VERSION : 0.1
   VAR
      _1s1 : Bool;
      _1s2 : Bool;
      _1s3 : Bool;
      _1s4 : Bool;
      _1s5 : Bool;
      _1s6 : Bool;
      _1s7 : Bool;
      _1s8 : Bool;
      _1s9 : Bool;
      _1s10 : Bool;
      _1sReserva2 : Bool;
      _1sReserva3 : Bool;
      _1sReserva4 : Bool;
      _1sReserva5 : Bool;
      _1sReserva6 : Bool;
      _1sReserva7 : Bool;
      _2s1 : Bool;
      _2s2 : Bool;
      _2s3 : Bool;
      _2s4 : Bool;
      _2s5 : Bool;
      _2s6 : Bool;
      _2s7 : Bool;
      _2s8 : Bool;
      _2s9 : Bool;
      _2s10 : Bool;
      _2sReserva2 : Bool;
      _2sReserva3 : Bool;
      _2sReserva4 : Bool;
      _2sReserva5 : Bool;
      _2sReserva6 : Bool;
      _2sReserva7 : Bool;
      _3s1 : Bool;
      _3s2 : Bool;
      _3s3 : Bool;
      _3s4 : Bool;
      _3s5 : Bool;
      _3s6 : Bool;
      _3s7 : Bool;
      _3s8 : Bool;
      _3s9 : Bool;
      _3s10 : Bool;
      _3Reserva2 : Bool;
      _3Reserva3 : Bool;
      _3Reserva4 : Bool;
      _3Reserva5 : Bool;
      _3Reserva6 : Bool;
      _3Reserva7 : Bool;
      _4s1 : Bool;
      _4s2 : Bool;
      _4s3 : Bool;
      _4s4 : Bool;
      _4s5 : Bool;
      _4s6 : Bool;
      _4s7 : Bool;
      _4s8 : Bool;
      _4s9 : Bool;
      _4s10 : Bool;
      _4sReserva2 : Bool;
      _4sReserva3 : Bool;
      _4sReserva4 : Bool;
      _4sReserva5 : Bool;
      _4sReserva6 : Bool;
      _4sReserva7 : Bool;
      _5s1 : Bool;
      _5s2 : Bool;
      _5s3 : Bool;
      _5s4 : Bool;
      _5s5 : Bool;
      _5s6 : Bool;
      _5s7 : Bool;
      _5s8 : Bool;
      _5s9 : Bool;
      _5s10 : Bool;
      _5sReserva2 : Bool;
      _5sReserva3 : Bool;
      _5sReserva4 : Bool;
      _5sReserva5 : Bool;
      _5sReserva6 : Bool;
      _5sReserva7 : Bool;
      _6s1 : Bool;
      _6s2 : Bool;
      _6s3 : Bool;
      _6s4 : Bool;
      _6s5 : Bool;
      _6s6 : Bool;
      _6s7 : Bool;
      _6s8 : Bool;
      _6s9 : Bool;
      _6s10 : Bool;
      _6sReserva2 : Bool;
      _6sReserva3 : Bool;
      _6sReserva4 : Bool;
      _6sReserva5 : Bool;
      _6sReserva6 : Bool;
      _6sReserva7 : Bool;
      _0s1 : Bool;   // No requiere Compresores
      _0s2 : Bool;   // Requiere 1 Compresor
      _0s3 : Bool;   // Requiere 2 Compresores
      _0s4 : Bool;   // Requiere 3 Compresores
      _0s5 : Bool;   // Requiere 4 Compresores
      _0s6 : Bool;   // Requiere 5 Compresores
      _0s7 : Bool;
      _0s8 : Bool;
      _0s9 : Bool;
      _0s10 : Bool;
      _0sReserva2 : Bool;
      _0sReserva3 : Bool;
      _0sReserva4 : Bool;
      _0sReserva5 : Bool;
      _0sReserva6 : Bool;
      _0sReserva7 : Bool;
   END_VAR
BEGIN
END_DATA_BLOCK

DATA_BLOCK "Concatenadoras"   // DB127
{ S7_Optimized_Access := 'FALSE' }
VERSION : 0.1
   VAR
      _1c1 : Bool;
      _1c2 : Bool;
      _1c3 : Bool;
      _1c4 : Bool;
      _1c5 : Bool;
      _1c6 : Bool;
      _1c7 : Bool;
      _1c8 : Bool;
      _1c9 : Bool;
      _1c10 : Bool;
      _1cReserva2 : Bool;
      _1cReserva3 : Bool;
      _1cReserva4 : Bool;
      _1cReserva5 : Bool;
      _1cReserva6 : Bool;
      _1cReserva7 : Bool;
      _2c1 : Bool;
      _2c2 : Bool;
      _2c3 : Bool;
      _2c4 : Bool;
      _2c5 : Bool;
      _2c6 : Bool;
      _2c7 : Bool;
      _2c8 : Bool;
      _2c9 : Bool;
      _2c10 : Bool;
      _2cReserva2 : Bool;
      _2cReserva3 : Bool;
      _2cReserva4 : Bool;
      _2cReserva5 : Bool;
      _2cReserva6 : Bool;
      _2cReserva7 : Bool;
      _3c1 : Bool;
      _3c2 : Bool;
      _3c3 : Bool;
      _3c4 : Bool;
      _3c5 : Bool;
      _3c6 : Bool;
      _3c7 : Bool;
      _3c8 : Bool;
      _3c9 : Bool;
      _3c10 : Bool;
      _3cReserva2 : Bool;
      _3cReserva3 : Bool;
      _3cReserva4 : Bool;
      _3cReserva5 : Bool;
      _3cReserva6 : Bool;
      _3cReserva7 : Bool;
      _4c1 : Bool;
      _4c2 : Bool;
      _4c3 : Bool;
      _4c4 : Bool;
      _4c5 : Bool;
      _4c6 : Bool;
      _4c7 : Bool;
      _4c8 : Bool;
      _4c9 : Bool;
      _4c10 : Bool;
      _4cReserva2 : Bool;
      _4cReserva3 : Bool;
      _4cReserva4 : Bool;
      _4cReserva5 : Bool;
      _4cReserva6 : Bool;
      _4cReserva7 : Bool;
      _5c1 : Bool;
      _5c2 : Bool;
      _5c3 : Bool;
      _5c4 : Bool;
      _5c5 : Bool;
      _5c6 : Bool;
      _5c7 : Bool;
      _5c8 : Bool;
      _5c9 : Bool;
      _5c10 : Bool;
      _5cReserva2 : Bool;
      _5cReserva3 : Bool;
      _5cReserva4 : Bool;
      _5cReserva5 : Bool;
      _5cReserva6 : Bool;
      _5cReserva7 : Bool;
      _6c1 : Bool;
      _6c2 : Bool;
      _6c3 : Bool;
      _6c4 : Bool;
      _6c5 : Bool;
      _6c6 : Bool;
      _6c7 : Bool;
      _6c8 : Bool;
      _6c9 : Bool;
      _6c10 : Bool;
      _6cReserva2 : Bool;
      _6cReserva3 : Bool;
      _6cReserva4 : Bool;
      _6cReserva5 : Bool;
      _6cReserva6 : Bool;
      _6cReserva7 : Bool;
      _0c1 : Bool;   // No requiere Compresores
      _0c2 : Bool;   // Requiere 1 Compresor
      _0c3 : Bool;   // Requiere 2 Compresores
      _0c4 : Bool;   // Requiere 3 Compresores
      _0c5 : Bool;   // Requiere 4 Compresores
      _0c6 : Bool;   // Requiere 5 Compresores
      _0c7 : Bool;
      _0c8 : Bool;
      _0c9 : Bool;
      _0c10 : Bool;
      _0cReserva2 : Bool;
      _0cReserva3 : Bool;
      _0cReserva4 : Bool;
      _0cReserva5 : Bool;
      _0cReserva6 : Bool;
      _0cReserva7 : Bool;
   END_VAR
BEGIN
END_DATA_BLOCK

DATA_BLOCK "Prioritarias"   // DB128
{ S7_Optimized_Access := 'FALSE' }
VERSION : 0.1
   VAR
      _1p1 : Bool;
      _1p2 : Bool;
      _1p3 : Bool;
      _1p4 : Bool;
      _1p5 : Bool;
      _1p6 : Bool;
      _1p7 : Bool;
      _1p8 : Bool;
      _1p9 : Bool;
      _1p10 : Bool;
      _1pReserva2 : Bool;
      _1pReserva3 : Bool;
      _1pReserva4 : Bool;
      _1pReserva5 : Bool;
      _1pReserva6 : Bool;
      _1pReserva7 : Bool;
      _2p1 : Bool;
      _2p2 : Bool;
      _2p3 : Bool;
      _2p4 : Bool;
      _2p5 : Bool;
      _2p6 : Bool;
      _2p7 : Bool;
      _2p8 : Bool;
      _2p9 : Bool;
      _2p10 : Bool;
      _2pReserva2 : Bool;
      _2pReserva3 : Bool;
      _2pReserva4 : Bool;
      _2pReserva5 : Bool;
      _2pReserva6 : Bool;
      _2pReserva7 : Bool;
      _3p1 : Bool;
      _3p2 : Bool;
      _3p3 : Bool;
      _3p4 : Bool;
      _3p5 : Bool;
      _3p6 : Bool;
      _3p7 : Bool;
      _3p8 : Bool;
      _3p9 : Bool;
      _3p10 : Bool;
      _3pReserva2 : Bool;
      _3pReserva3 : Bool;
      _3pReserva4 : Bool;
      _3pReserva5 : Bool;
      _3pReserva6 : Bool;
      _3pReserva7 : Bool;
      _4p1 : Bool;
      _4p2 : Bool;
      _4p3 : Bool;
      _4p4 : Bool;
      _4p5 : Bool;
      _4p6 : Bool;
      _4p7 : Bool;
      _4p8 : Bool;
      _4p9 : Bool;
      _4p10 : Bool;
      _4pReserva2 : Bool;
      _4pReserva3 : Bool;
      _4pReserva4 : Bool;
      _4pReserva5 : Bool;
      _4pReserva6 : Bool;
      _4pReserva7 : Bool;
      _5p1 : Bool;
      _5p2 : Bool;
      _5p3 : Bool;
      _5p4 : Bool;
      _5p5 : Bool;
      _5p6 : Bool;
      _5p7 : Bool;
      _5p8 : Bool;
      _5p9 : Bool;
      _5p10 : Bool;
      _5pReserva2 : Bool;
      _5pReserva3 : Bool;
      _5pReserva4 : Bool;
      _5pReserva5 : Bool;
      _5pReserva6 : Bool;
      _5pReserva7 : Bool;
      _6p1 : Bool;
      _6p2 : Bool;
      _6p3 : Bool;
      _6p4 : Bool;
      _6p5 : Bool;
      _6p6 : Bool;
      _6p7 : Bool;
      _6p8 : Bool;
      _6p9 : Bool;
      _6p10 : Bool;
      _6pReserva2 : Bool;
      _6pReserva3 : Bool;
      _6pReserva4 : Bool;
      _6pReserva5 : Bool;
      _6pReserva6 : Bool;
      _6pReserva7 : Bool;
      _0p1 : Bool;   // No requiere Compresores
      _0p2 : Bool;   // Requiere 1 Compresor
      _0p3 : Bool;   // Requiere 2 Compresores
      _0p4 : Bool;   // Requiere 3 Compresores
      _0p5 : Bool;   // Requiere 4 Compresores
      _0p6 : Bool;   // Requiere 5 Compresores
      _0p7 : Bool;
      _0p8 : Bool;
      _0p9 : Bool;
      _0p10 : Bool;
      _0pReserva2 : Bool;
      _0pReserva3 : Bool;
      _0pReserva4 : Bool;
      _0pReserva5 : Bool;
      _0pReserva6 : Bool;
      _0pReserva7 : Bool;
   END_VAR
BEGIN
END_DATA_BLOCK

DATA_BLOCK "FlancosMEst"   // DB129
{ S7_Optimized_Access := 'FALSE' }
VERSION : 0.1
   VAR
      fMan1 : Bool;   // flanco pasaje a modo manual
      fMan2 : Bool;   // flanco pasaje a modo manual
      fMan3 : Bool;   // flanco pasaje a modo manual
      fMan4 : Bool;   // flanco pasaje a modo manual
      fMan5 : Bool;   // flanco pasaje a modo manual
      fMan6 : Bool;
      fManP1 : Bool;   // Flanco selectora a manual prioridad 1
      fManP2 : Bool;   // Flanco selectora a manual prioridad 2
      fManP3 : Bool;   // Flanco selectora a manual prioridad 3
      fManP4 : Bool;   // Flanco selectora a manual prioridad 4
      fManP5 : Bool;   // Flanco selectora a manual prioridad 5
      fManP6 : Bool;
      fNoFal1 : Bool;   // flanco desapareció la falla Cmp 1
      fNoFal2 : Bool;   // flanco desapareció la falla Cmp 2
      fNoFal3 : Bool;   // flanco desapareció la falla Cmp 3
      fNoFal4 : Bool;   // flanco desapareció la falla Cmp 4
      fNoFal5 : Bool;   // flanco desapareció la falla Cmp 5
      fNoFal6 : Bool;
      fNoFaGen : Bool;   // fanco falla General
      fAlgCmpAuto : Bool;   // Flanco algún compresor pasó a automático
      ftSinReq1 : Bool;   // transición de compresor 1 sin requerimiento
      ftSinReq2 : Bool;   // transición de compresor 2 sin requerimiento
      ftSinReq3 : Bool;   // transición de compresor 3 sin requerimiento
      ftSinReq4 : Bool;   // transición de compresor 4 sin requerimiento
      ftSinReq5 : Bool;   // transición de compresor 5 sin requerimiento
      ftSinReq6 : Bool;
      ftSinReq : Bool;   // transición de algún compresor sin requerimiento
      fAut1 : Bool;   // Flanco automático compresor 1
      fAut2 : Bool;   // Flanco automático compresor 2
      fAut3 : Bool;   // Flanco automático compresor 3
      fAut4 : Bool;   // Flanco automático compresor 4
      fAut5 : Bool;   // Flanco automático compresor 5
      fAut6 : Bool;
      fNSop1 : Bool;   // Flanco negativo Sopladora 1
      fNSop2 : Bool;   // Flanco negativo Sopladora 2
      fNSop3 : Bool;   // Flanco negativo Sopladora 3
      fPSop1 : Bool;   // Flanco positivo Sopladora 1
      fPSop2 : Bool;   // Flanco positivo Sopladora 2
      fPSop3 : Bool;   // Flanco positivo Sopladora 3
   END_VAR
BEGIN
END_DATA_BLOCK

// folder: Compresores/Baja

DATA_BLOCK "PanelCompBAJA MTA"   // DB74
{ S7_Optimized_Access := 'FALSE' }
VERSION : 0.1
   VAR
      InhMC060 : Bool;   // Inhibición MC060
      InhMC061 : Bool;   // Inhibición MC061
      InhMC062 : Bool;   // Inhibición MC062
      InhMC063 : Bool;   // Inhibición MC063
      InhMC064 : Bool;   // Inhibición MC064
      InhMC065 : Bool;   // Inhibición MC065
      Flanco1MC060 : Bool;   // Flanco 1 MC060
      Flanco1MC061 : Bool;   // Flanco 1 MC061
      Flanco1MC062 : Bool;   // Flanco 1 MC062
      Flanco1MC063 : Bool;   // Flanco 1 MC063
      Flanco1MC064 : Bool;   // Flanco 1 MC064
      Flanco1MC065 : Bool;   // Flanco 1 MC065
      Flanco2MC060 : Bool;   // Flanco 2 MC060
      Flanco2MC061 : Bool;   // Flanco 2 MC061
      Flanco2MC062 : Bool;   // Flanco 2 MC062
      Flanco2MC063 : Bool;   // Flanco 2 MC063
      Flanco2MC064 : Bool;   // Flanco 2 MC064
      Flanco2MC065 : Bool;   // Flanco 2 MC065
      Flanco3MC060 : Bool;   // Flanco 3 MC060
      Flanco3MC061 : Bool;   // Flanco 3 MC061
      Flanco3MC062 : Bool;   // Flanco 3 MC062
      Flanco3MC063 : Bool;   // Flanco 3 MC063
      Flanco3MC064 : Bool;   // Flanco 3 MC064
      Flanco3MC065 : Bool;   // Flanco 3 MC065
      HabPanelMC060 : Bool;   // Habilitación desde Panel MC060
      HabPanelMC061 : Bool;   // Habilitación desde Panel MC061
      HabPanelMC062 : Bool;   // Habilitación desde Panel MC062
      HabPanelMC063 : Bool;   // Habilitación desde Panel MC063
      HabPanelMC064 : Bool;   // Habilitación desde Panel MC064
      HabPanelMC065 : Bool;   // Habilitación desde Panel MC065
      DeshabPanelMC060 : Bool;   // Deshabilitación desde Panel MC060
      DeshabPanelMC061 : Bool;   // Deshabilitación desde Panel MC061
      DeshabPanelMC062 : Bool;   // Deshabilitación desde Panel MC062
      DeshabPanelMC063 : Bool;   // Deshabilitación desde Panel MC063
      DeshabPanelMC064 : Bool;   // Deshabilitación desde Panel MC064
      DeshabPanelMC065 : Bool;   // Deshabilitación desde Panel MC065
      MarchaPanelMC060 : Bool;   // Marcha desde Panel MC060
      MarchaPanelMC061 : Bool;   // Marcha desde Panel MC061
      MarchaPanelMC062 : Bool;   // Marcha desde Panel MC062
      MarchaPanelMC063 : Bool;   // Marcha desde Panel MC063
      MarchaPanelMC064 : Bool;   // Marcha desde Panel MC064
      MarchaPanelMC065 : Bool;   // Marcha desde Panel MC065
      ParadaPanelMC060 : Bool;   // Parada desde Panel MC060
      ParadaPanelMC061 : Bool;   // Parada desde Panel MC061
      ParadaPanelMC062 : Bool;   // Parada desde Panel MC062
      ParadaPanelMC063 : Bool;   // Parada desde Panel MC063
      ParadaPanelMC064 : Bool;   // Parada desde Panel MC064
      ParadaPanelMC065 : Bool;   // Parada desde Panel MC065
      HabMC060 : Bool;   // Habilitado MC060
      HabMC061 : Bool;   // Habilitado MC061
      HabMC062 : Bool;   // Habilitado MC062
      HabMC063 : Bool;   // Habilitado MC063
      HabMC064 : Bool;   // Habilitado MC064
      HabMC065 : Bool;   // Habilitado MC065
      DeshabMC060 : Bool;   // Deshabilitado MC060
      DeshabMC061 : Bool;   // Deshabilitado MC061
      DeshabMC062 : Bool;   // Deshabilitado MC062
      DeshabMC063 : Bool;   // Deshabilitado MC063
      DeshabMC064 : Bool;   // Deshabilitado MC064
      DeshabMC065 : Bool;   // Deshabilitado MC065
      MarchaMC060 : Bool;   // Marchando MC060
      MarchaMC061 : Bool;   // Marchando MC061
      MarchaMC062 : Bool;   // Marchando MC062
      MarchaMC063 : Bool;   // Marchando MC063
      MarchaMC064 : Bool;   // Marchando MC064
      MarchaMC065 : Bool;   // Marchando MC065
      ParadaMC060 : Bool;   // Parando MC060
      ParadaMC061 : Bool;   // Parando MC061
      ParadaMC062 : Bool;   // Parando MC062
      ParadaMC063 : Bool;   // Parando MC063
      ParadaMC064 : Bool;   // Parando MC064
      ParadaMC065 : Bool;   // Parando MC065
      AnimMC060 : Byte;   // Animación MC060
      AnimMC061 : Byte;   // Animación MC061
      AnimMC062 : Byte;   // Animación MC062
      AnimMC063 : Byte;   // Animación MC063
      AnimMC064 : Byte;   // Animación MC064
      AnimMC065 : Byte;   // Animación MC065
      FallaGMTMC060 : Bool;   // Falla Térmica MC060
      FallaGMTMC061 : Bool;   // Falla Térmica MC061
      FallaGMTMC062 : Bool;   // Falla Térmica MC062
      FallaGMTMC063 : Bool;   // Falla Térmica MC063
      FallaGMTMC064 : Bool;   // Falla Térmica MC064
      FallaGMTMC065 : Bool;   // Falla Térmica MC065
      FallaCTCMC060 : Bool;   // Falla Contactor MC060
      FallaCTCMC061 : Bool;   // Falla Contactor MC061
      FallaCTCMC062 : Bool;   // Falla Contactor MC062
      FallaCTCMC063 : Bool;   // Falla Contactor MC063
      FallaCTCMC064 : Bool;   // Falla Contactor MC064
      FallaCTCMC065 : Bool;   // Falla Contactor MC065
      MantMC060 : Bool;   // Mantenimiento MC060
      MantMC061 : Bool;   // Mantenimiento MC061
      MantMC062 : Bool;   // Mantenimiento MC062
      MantMC063 : Bool;   // Mantenimiento MC063
      MantMC064 : Bool;   // Mantenimiento MC064
      MantMC065 : Bool;   // Mantenimiento MC065
      Reserva_1 : Bool;
      Reserva_11 : Bool;
      Reserva_12 : Bool;
      Reserva_13 : Bool;
      Reserva_14 : Bool;
      Reserva_15 : Bool;
      Reserva_16 : Bool;
      Reserva_17 : Bool;
      Reserva_18 : Bool;
      Reserva_19 : Bool;
      Reserva_110 : Bool;
      Reserva_111 : Bool;
      Reserva_112 : Bool;
      Reserva_113 : Bool;
      Reserva_114 : Bool;
      Reserva_115 : Bool;
      Reserva_116 : Bool;
      Reserva_117 : Bool;
      Reserva_118 : Bool;
      Reserva_119 : Bool;
      Reserva_120 : Bool;
      Reserva_121 : Bool;
      Reserva_122 : Bool;
      Reserva_123 : Bool;
      Reserva_124 : Bool;
      Reserva_125 : Bool;
      Reserva_126 : Bool;
      Reserva_127 : Bool;
      Reserva_128 : Bool;
      Reserva_129 : Bool;
      Reserva_130 : Bool;
      Reserva_131 : Bool;
      Reserva_132 : Bool;
      Reserva_133 : Bool;
      Reserva_134 : Bool;
      Reserva_135 : Bool;
      Reserva_136 : Bool;
      Reserva_137 : Bool;
      Reserva_138 : Bool;
      Reserva_139 : Bool;
      Reserva_140 : Bool;
      Reserva_141 : Bool;
      Reserva_142 : Bool;
      Reserva_143 : Bool;
   END_VAR
BEGIN
END_DATA_BLOCK

DATA_BLOCK "CmpBajaAuto"   // DB93
{ S7_Optimized_Access := 'FALSE' }
VERSION : 0.1
   VAR
      AutoMC060 : Bool;   // MC060 en modo auto
      AutoMC061 : Bool;   // MC061 en modo auto
      AutoMC062 : Bool;   // MC062 en modo auto
      AutoMC063 : Bool;   // MC063 en modo auto
      AutoMC064 : Bool;   // MC064 en modo auto
      SPonMC060 : Real;   // SetPoint de arranque MC060
      SPonMC061 : Real;   // SetPoint de arranque MC061
      SPonMC062 : Real;   // SetPoint de arranque MC062
      SPonMC063 : Real;   // SetPoint de arranque MC063
      SPonMC064 : Real;   // SetPoint de arranque MC064
      SPoffMC060 : Real;   // SetPoint de Parada MC060
      SPoffMC061 : Real;   // SetPoint de Parada MC061
      SPoffMC062 : Real;   // SetPoint de Parada MC062
      SPoffMC063 : Real;   // SetPoint de Parada MC063
      SPoffMC064 : Real;   // SetPoint de Parada MC064
      AutoArrMC060 : Bool;   // Arranque automático MC060
      AutoArrMC061 : Bool;   // Arranque automático MC061
      AutoArrMC062 : Bool;   // Arranque automático MC062
      AutoArrMC063 : Bool;   // Arranque automático MC063
      AutoArrMC064 : Bool;   // Arranque automático MC064
      AutoArrEfMC060 : Bool;   // Arranque automático efectivo MC060
      AutoArrEfMC061 : Bool;   // Arranque automático efectivo MC061
      AutoArrEfMC062 : Bool;   // Arranque automático efectivo MC062
      AutoArrEfMC063 : Bool;   // Arranque automático efectivo MC063
      AutoArrEfMC064 : Bool;   // Arranque automático efectivo MC064
      MenuMC060 : Int;   // Byte animación para menú MC060
      MenuMC061 : Int;   // Byte animación para menú MC061
      MenuMC062 : Int;   // Byte animación para menú MC062
      MenuMC063 : Int;   // Byte animación para menú MC063
      MenuMC064 : Int;   // Byte animación para menú MC064
   END_VAR
BEGIN
END_DATA_BLOCK

// folder: Entradas Analógicas

DATA_BLOCK "CaudalPotencia"   // DB26
{ S7_Optimized_Access := 'FALSE' }
VERSION : 0.1
   VAR
      lecCaudal : Real := 0.0;
      lecPotencia : Real := 0.0;
      HI_caudal : Real := 100.0;
      LO_caudal : Real := 0.0;
      HI_potencia : Real := 100.0;
      LO_potencia : Real := 0.0;
   END_VAR
BEGIN
END_DATA_BLOCK

DATA_BLOCK "LectAnalógicasMTA"   // DB52
{ S7_Optimized_Access := 'FALSE' }
VERSION : 0.1
   VAR
      TempCav : Real;   // Temperatura torres cavaleto
      TempChill : Real;   // Temperatura torres chillers
      PresAlta1 : Real;   // Presión de Alta 1
      PresAlta12 : Real;   // Presión de Alta 2
      PresBaja : Real;   // Presión de Baja
      PreAltaHH : Real;   // Presión de Alta Muy Alta
      PreAltaH : Real;   // Presión de Alta Alta
      PreAltaL : Real;   // Presión de Alta Baja
      PreAltaLL : Real;   // Presión de Alta Muy Baja
      PreBajaHH : Real;   // Presión de Baja Muy Alta
      PreBajaH : Real;   // Presión de Baja Alta
      PreBajaL : Real;   // Presión de Baja Baja
      PreBajaLL : Real;   // Presión de Baja Muy Baja
      PresionALTA : Real;   // Presión de Alta Final
   END_VAR
BEGIN
END_DATA_BLOCK

DATA_BLOCK "EntradasAnalógicas MTA"   // DB72
{ S7_Optimized_Access := 'FALSE' }
VERSION : 0.1
   VAR
      PresAire : Real;
      TempTanque1CH : Real;
      TempTanque2CH : Real;
      TempTorresCH : Real;
      FallaAIRE : Bool;
      FallaTanque1 : Bool;
      FallaTanque2 : Bool;
      FallaTorres : Bool;
   END_VAR
BEGIN
END_DATA_BLOCK

// folder: Horas de Marcha

DATA_BLOCK "Varios"   // DB2
{ S7_Optimized_Access := 'FALSE' }
VERSION : 0.1
   VAR
      HorasMantMC001_1 : DInt := 8000;   // Cantidad de Horas Máxima para un compresor
      HorasMantMC002_1 : DInt := 8000;
      HorasMantMC003_1 : DInt := 10005;
      HorasMantMC004_1 : DInt := 8000;
      HorasMantMC005_1 : DInt := 8000;
      HorasMantMC006_1 : DInt := 8000;
      HorasMantMC001_2 : DInt := 999999;
      HorasMantMC002_2 : DInt := 999999;
      HorasMantMC003_2 : DInt := 10013;
      HorasMantMC004_2 : DInt := 999999;
      HorasMantMC005_2 : DInt := 999999;
      HorasMantMC006_2 : DInt := 999999;
      UltimoMantMC001_1 : DInt := 90120;
      UltimoMantMC002_1 : DInt := 19431;
      UltimoMantMC003_1 : DInt := 0;
      UltimoMantMC004_1 : DInt := 65362;
      UltimoMantMC005_1 : DInt := 96802;
      UltimoMantMC006_1 : DInt := 0;
      UltimoMantMC001_2 : DInt := 0;
      UltimoMantMC002_2 : DInt := 0;
      UltimoMantMC003_2 : DInt := 0;
      UltimoMantMC004_2 : DInt := 0;
      UltimoMantMC005_2 : DInt := 0;
      UltimoMantMC006_2 : DInt := 3324;
      HorasMantMS050 : DInt := 8000;
      HorasMantMS051 : DInt := 10007;
      HorasMantMS052 : DInt := 10014;
      HorasMantMS053 : DInt := 10015;
      UltimoMantMS050 : DInt := 0;
      UltimoMantMS051 : DInt := 0;
      UltimoMantMS052 : DInt := 0;
      UltimoMantMS053 : DInt := 0;
      HorasMantMC060_1 : DInt := 2000;
      HorasMantMC061_1 : DInt := 2000;
      HorasMantMC062_1 : DInt := 1;
      HorasMantMC063_1 : DInt := 2000;
      HorasMantMC064_1 : DInt := 1;
      HorasMantMC065_1 : DInt := 0;
      HorasMantMC060_2 : DInt := 4000;
      HorasMantMC061_2 : DInt := 4000;
      HorasMantMC062_2 : DInt := 1;
      HorasMantMC063_2 : DInt := 4000;
      HorasMantMC064_2 : DInt := 1;
      HorasMantMC065_2 : DInt := 0;
      HorasMantMC060_3 : DInt := 8000;
      HorasMantMC061_3 : DInt := 8000;
      HorasMantMC062_3 : DInt := 1;
      HorasMantMC063_3 : DInt := 8000;
      HorasMantMC064_3 : DInt := 1;
      HorasMantMC065_3 : DInt := 0;
      HorasMantMC060_4 : DInt := 20000;
      HorasMantMC061_4 : DInt := 80000;
      HorasMantMC062_4 : DInt := 1;
      HorasMantMC063_4 : DInt := 24000;
      HorasMantMC064_4 : DInt := 1;
      HorasMantMC065_4 : DInt := 0;
      HorasMantMC060_5 : DInt := 0;
      HorasMantMC061_5 : DInt := 80000;
      HorasMantMC062_5 : DInt := 1;
      HorasMantMC063_5 : DInt := 0;
      HorasMantMC064_5 : DInt := 1;
      HorasMantMC065_5 : DInt := 0;
      UltimoMantMC060_1 : DInt := 5643;
      UltimoMantMC061_1 : DInt := 38265;
      UltimoMantMC062_1 : DInt := 0;
      UltimoMantMC063_1 : DInt := 37701;
      UltimoMantMC064_1 : DInt := 0;
      UltimoMantMC065_1 : DInt := 0;
      UltimoMantMC060_2 : DInt := 5643;
      UltimoMantMC061_2 : DInt := 38265;
      UltimoMantMC062_2 : DInt := 0;
      UltimoMantMC063_2 : DInt := 37701;
      UltimoMantMC064_2 : DInt := 0;
      UltimoMantMC065_2 : DInt := 0;
      UltimoMantMC060_3 : DInt := 5643;
      UltimoMantMC061_3 : DInt := 38265;
      UltimoMantMC062_3 : DInt := 0;
      UltimoMantMC063_3 : DInt := 30970;
      UltimoMantMC064_3 : DInt := 0;
      UltimoMantMC065_3 : DInt := 0;
      UltimoMantMC060_4 : DInt := 0;
      UltimoMantMC061_4 : DInt := 0;
      UltimoMantMC062_4 : DInt := 0;
      UltimoMantMC063_4 : DInt := 30970;
      UltimoMantMC064_4 : DInt := 0;
      UltimoMantMC065_4 : DInt := 0;
      UltimoMantMC060_5 : DInt := 40000;
      UltimoMantMC061_5 : DInt := 0;
      UltimoMantMC062_5 : DInt := 0;
      UltimoMantMC063_5 : DInt := 0;
      UltimoMantMC064_5 : DInt := 0;
      UltimoMantMC065_5 : DInt := 0;
      HorasMantMS054_1 : DInt := 7000;
      HorasMantMS055_1 : DInt := 0;
      HorasMantMS056_1 : DInt := 0;
      HorasMantMS054_2 : DInt := 7001;
      HorasMantMS055_2 : DInt := 7003;
      HorasMantMS056_2 : DInt := 0;
      UltimoMantMS054_1 : DInt := 0;
      UltimoMantMS055_1 : DInt := 7002;
      UltimoMantMS056_1 : DInt := 0;
      UltimoMantMS054_2 : DInt := 0;
      UltimoMantMS055_2 : DInt := 0;
      UltimoMantMS056_2 : DInt := 0;
      HorasMantBost1 : DInt := 15000;
      HorasMantBost2 : DInt := 15000;
      UltimoMantBoost1 : DInt := 0;
      UltimoMantBoost2 : DInt := 0;
   END_VAR
BEGIN
END_DATA_BLOCK

DATA_BLOCK "HorasSecAlta"   // DB19
{ S7_Optimized_Access := 'FALSE' }
VERSION : 0.1
   VAR
      HMMS050 : DInt;
      HMMS051 : DInt;
      HMMS052 : DInt;
      HMMS053 : DInt;
      MMMS050 : Int;
      MMMS051 : Int;
      MMMS052 : Int;
      MMMS053 : Int;
      SMMS050 : Int;
      SMMS051 : Int;
      SMMS052 : Int;
      SMMS053 : Int;
   END_VAR
BEGIN
END_DATA_BLOCK

DATA_BLOCK "HorasCmpBaja"   // DB20
{ S7_Optimized_Access := 'FALSE' }
VERSION : 0.1
   VAR
      HMMC060 : DInt;
      HMMC061 : DInt;
      HMMC062 : DInt;
      HMMC063 : DInt;
      HMMC064 : DInt;
      HMMC065 : DInt;
      MMMC060 : Int;
      MMMC061 : Int;
      MMMC062 : Int;
      MMMC063 : Int;
      MMMC064 : Int;
      MMMC065 : Int;
      SMMC060 : Int;
      SMMC061 : Int;
      SMMC062 : Int;
      SMMC063 : Int;
      SMMC064 : Int;
      SMMC065 : Int;
   END_VAR
BEGIN
END_DATA_BLOCK

DATA_BLOCK "HorasSecBaja"   // DB24
{ S7_Optimized_Access := 'FALSE' }
VERSION : 0.1
   VAR
      HMMS054 : DInt;
      HMMS055 : DInt;
      HMMS056 : DInt;
      MMMS054 : Int;
      MMMS055 : Int;
      MMMS056 : Int;
      SMMS054 : Int;
      SMMS055 : Int;
      SMMS056 : Int;
   END_VAR
BEGIN
END_DATA_BLOCK

DATA_BLOCK "SumaOB35 MTA"   // DB73
{ S7_Optimized_Access := 'FALSE' }
VERSION : 0.1
   VAR
      HMMC001 : DInt;   // Horas acumuladas compresor 1
      HMMC002 : DInt;   // Horas acumuladas compresor 2
      HMMC003 : DInt;   // Horas acumuladas compresor 3
      HMMC004 : DInt;   // Horas acumuladas compresor 4
      HMMC005 : DInt;   // Horas acumuladas compresor 5
      HMMC006 : DInt;
      MMMC001 : Int;   // Minutos acumuladas compresor 1
      MMMC002 : Int;   // Minutos acumuladas compresor 2
      MMMC003 : Int;   // Minutos acumuladas compresor 3
      MMMC004 : Int;   // Minutos acumuladas compresor 4
      MMMC005 : Int;   // Minutos acumuladas compresor 5
      MMMC006 : Int;
      PrioridadArranqueMC001 : Int;
      PrioridadArranqueMC002 : Int;
      PrioridadArranqueMC003 : Int;
      PrioridadArranqueMC004 : Int;
      PrioridadArranqueMC005 : Int;
      PrioridadArranqueMC006 : Int;
      PrioridadParadaMC001 : Int;
      PrioridadParadaMC002 : Int;
      PrioridadParadaMC003 : Int;
      PrioridadParadaMC004 : Int;
      PrioridadParadaMC005 : Int;
      PrioridadParadaMC006 : Int;
      HorasMin : DInt;
      HorasMax : DInt;
      MotoreEnMarcha : Int;
      SMMC001 : Int;   // Segundos acumuladas compresor 1
      SMMC002 : Int;   // Segundos acumuladas compresor 2
      SMMC003 : Int;   // Segundos acumuladas compresor 3
      SMMC004 : Int;   // Segundos acumuladas compresor 4
      SMMC005 : Int;   // Segundos acumuladas compresor 5
      SMMC006 : Int;
      ByteMotoresEnAUTO : Byte;
      ByteMotoresEnMarcha : Byte;
   END_VAR
BEGIN
END_DATA_BLOCK

// folder: Panel

DATA_BLOCK "Bloque de animacion MTA"   // DB46
{ S7_Optimized_Access := 'FALSE' }
VERSION : 0.1
   VAR
      AnimacionMP010 : Byte;
      AnimacionMP011 : Byte;
      AnimacionMP012 : Byte;
      AnimacionMP013 : Byte;
      AnimacionMP018 : Byte;
      AnimacionMP019 : Byte;
      AnimacionMT007 : Byte;
      AnimacionMT008 : Byte;
      AnimacionMT009 : Byte;
      AnimacionMT010 : Byte;
      AnimacionV001 : Byte;
      AnimacionV002 : Byte;
      AnimacionV003 : Byte;
      MenuMS050 : Int;   // Byte animación para menú MS050
      MenuMS051 : Int;   // Byte animación para menú MS051
      MenuMS052 : Int;   // Byte animación para menú MS052
      MenuMS053 : Int;   // Byte animación para menú MS053
      MenuMS054 : Int;   // Byte animación para menú MS054
      MenuV001 : Int;   // Byte animación para menú V001
      MenuV002 : Int;   // Byte animación para menú V002
      MenuV003 : Int;   // Byte animación para menú V003
      AnimacionMS054 : Byte;
      AnimacionMS055 : Byte;
      MenuV030 : Int;   // Byte animación para menú V030
      MenuV031 : Int;   // Byte animación para menú V031
      AnimMV030 : Byte;   // Animación MV030
      AnimMV031 : Byte;   // Animación MV031
      AnimMP014 : Byte;   // Animación MP014
      AnimMP015 : Byte;   // Animación MP015
      AnimMC001 : Byte;   // Animación MC001
      AnimMC002 : Byte;   // Animación MC002
      AnimMC003 : Byte;   // Animación MC003
      AnimMC004 : Byte;   // Animación MC004
      AnimMC005 : Byte;   // Animación MC005
      AnimMC006 : Byte;
      Reserva17 : Byte;
      Reserva18 : Byte;
      Reserva19 : Byte;
      Reserva20 : Byte;
      Reserva21 : Byte;
      Reserva22 : Byte;
      Reserva23 : Byte;
      Reserva24 : Byte;
      Reserva25 : Byte;
      Reserva26 : Byte;
      Reserva27 : Byte;
      Reserva28 : Byte;
      Reserva29 : Byte;
      Reserva30 : Byte;
      Reserva31 : Byte;
      Reserva32 : Byte;
      Reserva33 : Byte;
      Reserva34 : Byte;
      Reserva35 : Byte;
      Reserva36 : Byte;
      Reserva37 : Byte;
      Reserva38 : Byte;
      Reserva39 : Byte;
      Reserva40 : Byte;
      Reserva41 : Byte;
      Reserva42 : Byte;
      Reserva43 : Byte;
      Reserva44 : Byte;
      Reserva45 : Byte;
      Reserva46 : Byte;
      Reserva47 : Byte;
      Reserva48 : Byte;
      Reserva49 : Byte;
      Reserva50 : Byte;
      Reserva51 : Byte;
      Reserva52 : Byte;
      Reserva53 : Byte;
      Reserva54 : Byte;
      Reserva55 : Byte;
      Reserva56 : Byte;
      Reserva57 : Byte;
      Reserva58 : Byte;
      Reserva59 : Byte;
      Reserva60 : Byte;
      Reserva61 : Byte;
      Reserva62 : Byte;
      Reserva63 : Byte;
      Reserva64 : Byte;
      Reserva65 : Byte;
      Reserva66 : Byte;
      Reserva67 : Byte;
      Reserva68 : Byte;
      Reserva69 : Byte;
      Reserva70 : Byte;
      Reserva71 : Byte;
      Reserva72 : Byte;
      Reserva73 : Byte;
      Reserva74 : Byte;
   END_VAR
BEGIN
END_DATA_BLOCK

DATA_BLOCK "PanelMotChillMTA"   // DB90
{ S7_Optimized_Access := 'FALSE' }
VERSION : 0.1
   VAR
      InhMT007 : Bool;   // Inhibición MT007
      InhMT008 : Bool;   // Inhibición MT008
      InhMT009 : Bool;   // Inhibición MT009
      InhMT010 : Bool;   // Inhibición MT010
      InhMP010 : Bool;   // Inhibición MP010
      InhMP011 : Bool;   // Inhibición MP011
      InhMP012 : Bool;   // Inhibición MP012
      InhMP013 : Bool;   // Inhibición MP013
      InhMP018 : Bool;   // Inhibición MP018
      InhMP019 : Bool;   // Inhibición MP019
      InhV001 : Bool;   // Inhibición V001
      InhV002 : Bool;   // Inhibición V002
      InhV003 : Bool;   // Inhibición V003
      Flanco1MT007 : Bool;   // Flanco 1 MT007
      Flanco1MT008 : Bool;   // Flanco 1 MT008
      Flanco1MT009 : Bool;   // Flanco 1 MT009
      Flanco1MT010 : Bool;   // Flanco 1 MT010
      Flanco1MP010 : Bool;   // Flanco 1 MP010
      Flanco1MP011 : Bool;   // Flanco 1 MP011
      Flanco1MP012 : Bool;   // Flanco 1 MP012
      Flanco1MP013 : Bool;   // Flanco 1 MP013
      Flanco1MP018 : Bool;   // Flanco 1 MP018
      Flanco1MP019 : Bool;   // Flanco 1 MP019
      Flanco1V001 : Bool;   // Flanco 1 V001
      Flanco1V002 : Bool;   // Flanco 1 V002
      Flanco1V003 : Bool;   // Flanco 1 V003
      Flanco2MT007 : Bool;   // Flanco 2 MT007
      Flanco2MT008 : Bool;   // Flanco 2 MT008
      Flanco2MT009 : Bool;   // Flanco 2 MT009
      Flanco2MT010 : Bool;   // Flanco 2 MT010
      Flanco2MP010 : Bool;   // Flanco 2 MP010
      Flanco2MP011 : Bool;   // Flanco 2 MP011
      Flanco2MP012 : Bool;   // Flanco 2 MP012
      Flanco2MP013 : Bool;   // Flanco 2 MP013
      Flanco2MP018 : Bool;   // Flanco 2 MP018
      Flanco2MP019 : Bool;   // Flanco 2 MP019
      Flanco2V001 : Bool;   // Flanco 2 V001
      Flanco2V002 : Bool;   // Flanco 2 V002
      Flanco2V003 : Bool;   // Flanco 2 V003
      Flanco3MT007 : Bool;   // Flanco 3 MT007
      Flanco3MT008 : Bool;   // Flanco 3 MT008
      Flanco3MT009 : Bool;   // Flanco 3 MT009
      Flanco3MT010 : Bool;   // Flanco 3 MT010
      Flanco3MP010 : Bool;   // Flanco 3 MP010
      Flanco3MP011 : Bool;   // Flanco 3 MP011
      Flanco3MP012 : Bool;   // Flanco 3 MP012
      Flanco3MP013 : Bool;   // Flanco 3 MP013
      Flanco3MP018 : Bool;   // Flanco 3 MP018
      Flanco3MP019 : Bool;   // Flanco 3 MP019
      Flanco3V001 : Bool;   // Flanco 3 V001
      Flanco3V002 : Bool;   // Flanco 3 V002
      Flanco3V003 : Bool;   // Flanco 3 V003
      HabPanelMT007 : Bool;   // Habilitación desde Panel MT007
      HabPanelMT008 : Bool;   // Habilitación desde Panel MT008
      HabPanelMT009 : Bool;   // Habilitación desde Panel MT009
      HabPanelMT010 : Bool;   // Habilitación desde Panel MT010
      HabPanelMP010 : Bool;   // Habilitación desde Panel MP010
      HabPanelMP011 : Bool;   // Habilitación desde Panel MP011
      HabPanelMP012 : Bool;   // Habilitación desde Panel MP012
      HabPanelMP013 : Bool;   // Habilitación desde Panel MP013
      HabPanelMP018 : Bool;   // Habilitación desde Panel MP018
      HabPanelMP019 : Bool;   // Habilitación desde Panel MP019
      HabPanelV001 : Bool;   // Habilitación desde Panel V001
      HabPanelV002 : Bool;   // Habilitación desde Panel V002
      HabPanelV003 : Bool;   // Habilitación desde Panel V003
      DeshabPanelMT007 : Bool;   // Deshabilitación desde Panel MT007
      DeshabPanelMT008 : Bool;   // Deshabilitación desde Panel MT008
      DeshabPanelMT009 : Bool;   // Deshabilitación desde Panel MT009
      DeshabPanelMT010 : Bool;   // Deshabilitación desde Panel MT010
      DeshabPanelMP010 : Bool;   // Deshabilitación desde Panel MP010
      DeshabPanelMP011 : Bool;   // Deshabilitación desde Panel MP011
      DeshabPanelMP012 : Bool;   // Deshabilitación desde Panel MP012
      DeshabPanelMP013 : Bool;   // Deshabilitación desde Panel MP013
      DeshabPanelMP018 : Bool;   // Deshabilitación desde Panel MP018
      DeshabPanelMP019 : Bool;   // Deshabilitación desde Panel MP019
      DeshabPanelV001 : Bool;   // Deshabilitación desde Panel V001
      DeshabPanelV002 : Bool;   // Deshabilitación desde Panel V002
      DeshabPanelV003 : Bool;   // Deshabilitación desde Panel V003
      MarchaPanelMT007 : Bool;   // Marcha desde Panel MT007
      MarchaPanelMT008 : Bool;   // Marcha desde Panel MT008
      MarchaPanelMT009 : Bool;   // Marcha desde Panel MT009
      MarchaPanelMT010 : Bool;   // Marcha desde Panel MT010
      MarchaPanelMP010 : Bool;   // Marcha desde Panel MP010
      MarchaPanelMP011 : Bool;   // Marcha desde Panel MP011
      MarchaPanelMP012 : Bool;   // Marcha desde Panel MP012
      MarchaPanelMP013 : Bool;   // Marcha desde Panel MP013
      MarchaPanelMP018 : Bool;   // Marcha desde Panel MP018
      MarchaPanelMP019 : Bool;   // Marcha desde Panel MP019
      MarchaPanelV001 : Bool;   // Marcha desde Panel V001
      MarchaPanelV002 : Bool;   // Marcha desde Panel V002
      MarchaPanelV003 : Bool;   // Marcha desde Panel V003
      ParadaPanelMT007 : Bool;   // Parada desde Panel MT007
      ParadaPanelMT008 : Bool;   // Parada desde Panel MT008
      ParadaPanelMT009 : Bool;   // Parada desde Panel MT009
      ParadaPanelMT010 : Bool;   // Parada desde Panel MT010
      ParadaPanelMP010 : Bool;   // Parada desde Panel MP010
      ParadaPanelMP011 : Bool;   // Parada desde Panel MP011
      ParadaPanelMP012 : Bool;   // Parada desde Panel MP012
      ParadaPanelMP013 : Bool;   // Parada desde Panel MP013
      ParadaPanelMP018 : Bool;   // Parada desde Panel MP018
      ParadaPanelMP019 : Bool;   // Parada desde Panel MP019
      ParadaPanelV001 : Bool;   // Parada desde Panel V001
      ParadaPanelV002 : Bool;   // Parada desde Panel V002
      ParadaPanelV003 : Bool;   // Parada desde Panel V003
      HabMT007 : Bool;   // Habilitado MT007
      HabMT008 : Bool := TRUE;   // Habilitado MT008
      HabMT009 : Bool;   // Habilitado MT009
      HabMT010 : Bool;   // Habilitado MT010
      HabMP010 : Bool;   // Habilitado MP010
      HabMP011 : Bool := TRUE;   // Habilitado MP011
      HabMP012 : Bool;   // Habilitado MP012
      HabMP013 : Bool;   // Habilitado MP013
      HabMP018 : Bool := TRUE;   // Habilitado MP018
      HabMP019 : Bool;   // Habilitado MP019
      HabV001 : Bool;   // Habilitado V001
      HabV002 : Bool;   // Habilitado V002
      HabV003 : Bool;   // Habilitado V003
      DeshabMT007 : Bool;   // Deshabilitado MT007
      DeshabMT008 : Bool;   // Deshabilitado MT008
      DeshabMT009 : Bool;   // Deshabilitado MT009
      DeshabMT010 : Bool;   // Deshabilitado MT010
      DeshabMP010 : Bool;   // Deshabilitado MP010
      DeshabMP011 : Bool;   // Deshabilitado MP011
      DeshabMP012 : Bool;   // Deshabilitado MP012
      DeshabMP013 : Bool;   // Deshabilitado MP013
      DeshabMP018 : Bool;   // Deshabilitado MP018
      DeshabMP019 : Bool;   // Deshabilitado MP019
      DeshabV001 : Bool;   // Deshabilitado V001
      DeshabV002 : Bool;   // Deshabilitado V002
      DeshabV003 : Bool;   // Deshabilitado V003
      MarchaMT007 : Bool;   // Marchando MT007
      MarchaMT008 : Bool := TRUE;   // Marchando MT008
      MarchaMT009 : Bool;   // Marchando MT009
      MarchaMT010 : Bool;   // Marchando MT010
      MarchaMP010 : Bool;   // Marchando MP010
      MarchaMP011 : Bool := TRUE;   // Marchando MP011
      MarchaMP012 : Bool;   // Marchando MP012
      MarchaMP013 : Bool;   // Marchando MP013
      MarchaMP018 : Bool := TRUE;   // Marchando MP018
      MarchaMP019 : Bool;   // Marchando MP019
      MarchaV001 : Bool;   // Marchando V001
      MarchaV002 : Bool;   // Marchando V002
      MarchaV003 : Bool;   // Marchando V003
      ParadaMT007 : Bool;   // Parando MT007
      ParadaMT008 : Bool;   // Parando MT008
      ParadaMT009 : Bool;   // Parando MT009
      ParadaMT010 : Bool;   // Parando MT010
      ParadaMP010 : Bool;   // Parando MP010
      ParadaMP011 : Bool;   // Parando MP011
      ParadaMP012 : Bool;   // Parando MP012
      ParadaMP013 : Bool;   // Parando MP013
      ParadaMP018 : Bool;   // Parando MP018
      ParadaMP019 : Bool;   // Parando MP019
      ParadaV001 : Bool;   // Parando V001
      ParadaV002 : Bool;   // Parando V002
      ParadaV003 : Bool;   // Parando V003
      AnimMT007 : Byte;   // Animación MT007
      AnimMT008 : Byte;   // Animación MT008
      AnimMT009 : Byte;   // Animación MT009
      AnimMT010 : Byte;   // Animación MT010
      AnimMP010 : Byte;   // Animación MP010
      AnimMP011 : Byte;   // Animación MP011
      AnimMP012 : Byte;   // Animación MP012
      AnimMP013 : Byte;   // Animación MP013
      AnimMP018 : Byte;   // Animación MP018
      AnimMP019 : Byte;   // Animación MP019
      AnimV001 : Byte;   // Animación V001
      AnimV002 : Byte;   // Animación V002
      AnimV003 : Byte;   // Animación V003
      Reserva_1 : Bool;
      Reserva_11 : Bool;
      Reserva_12 : Bool;
      Reserva_13 : Bool;
      Reserva_14 : Bool;
      Reserva_15 : Bool;
      Reserva_16 : Bool;
      Reserva_17 : Bool;
      Reserva_18 : Bool;
      Reserva_19 : Bool;
      Reserva_110 : Bool;
      Reserva_111 : Bool;
      Reserva_112 : Bool;
      Reserva_113 : Bool;
      Reserva_114 : Bool;
      Reserva_115 : Bool;
      Reserva_116 : Bool;
      Reserva_117 : Bool;
      Reserva_118 : Bool;
      Reserva_119 : Bool;
      Reserva_120 : Bool;
      Reserva_121 : Bool;
      Reserva_122 : Bool;
      Reserva_123 : Bool;
      Reserva_124 : Bool;
      Reserva_125 : Bool;
      Reserva_126 : Bool;
      Reserva_127 : Bool;
      Reserva_128 : Bool;
      Reserva_129 : Bool;
      Reserva_130 : Bool;
      Reserva_131 : Bool;
      Reserva_132 : Bool;
      Reserva_133 : Bool;
      Reserva_134 : Bool;
      Reserva_135 : Bool;
      Reserva_136 : Bool;
      Reserva_137 : Bool;
      Reserva_138 : Bool;
      Reserva_139 : Bool;
      Reserva_140 : Bool;
      Reserva_141 : Bool;
      Reserva_142 : Bool;
      Reserva_143 : Bool;
   END_VAR
BEGIN
END_DATA_BLOCK

// folder: Panel/Iluminación

DATA_BLOCK "DBIluminaciónMTA"   // DB87
{ S7_Optimized_Access := 'FALSE' }
VERSION : 0.1
   VAR
      TiempoDeEncendido : Word;
      EncendidoPanel : Bool;
      ApagadoPanel : Bool;
      Encendido : Bool;
      MantenerEncendida : Bool;
      AuxiliarEncendidoPermane : Bool;
      FLANCOP : Bool;
      FLANCON : Bool;
      EcendidoPLS : Bool;
      ApagadoPLS : Bool;
      TiempoPANEL : S5Time;
      AuxiliarCalculo : Int;
      TiempoPANEL1 : S5Time;
   END_VAR
BEGIN
END_DATA_BLOCK

// folder: Secadores/Alta

DATA_BLOCK "PanelSecALTA"   // DB81
{ S7_Optimized_Access := 'FALSE' }
VERSION : 0.1
   VAR
      InhMS050 : Bool;   // Inhibición MS050
      InhMS051 : Bool;   // Inhibición MS051
      InhMS052 : Bool;   // Inhibición MS052
      InhMS053 : Bool;   // Inhibición MS053
      Flanco1MS050 : Bool;   // Flanco 1 MS050
      Flanco1MS051 : Bool;   // Flanco 1 MS051
      Flanco1MS052 : Bool;   // Flanco 1 MS052
      Flanco1MS053 : Bool;   // Flanco 1 MS053
      Flanco2MS050 : Bool;   // Flanco 2 MS050
      Flanco2MS051 : Bool;   // Flanco 2 MS051
      Flanco2MS052 : Bool;   // Flanco 2 MS052
      Flanco2MS053 : Bool;   // Flanco 2 MS053
      Flanco3MS050 : Bool;   // Flanco 3 MS050
      Flanco3MS051 : Bool;   // Flanco 3 MS051
      Flanco3MS052 : Bool;   // Flanco 3 MS052
      Flanco3MS053 : Bool;   // Flanco 3 MS053
      HabPanelMS050 : Bool;   // Habilitación desde Panel MS050
      HabPanelMS051 : Bool;   // Habilitación desde Panel MS051
      HabPanelMS052 : Bool;   // Habilitación desde Panel MS052
      HabPanelMS053 : Bool;   // Habilitación desde Panel MS053
      DeshabPanelMS050 : Bool;   // Deshabilitación desde Panel MS050
      DeshabPanelMS051 : Bool;   // Deshabilitación desde Panel MS051
      DeshabPanelMS052 : Bool;   // Deshabilitación desde Panel MS052
      DeshabPanelMS053 : Bool;   // Deshabilitación desde Panel MS053
      MarchaPanelMS050 : Bool;   // Marcha desde Panel MS050
      MarchaPanelMS051 : Bool;   // Marcha desde Panel MS051
      MarchaPanelMS052 : Bool;   // Marcha desde Panel MS052
      MarchaPanelMS053 : Bool;   // Marcha desde Panel MS053
      ParadaPanelMS050 : Bool;   // Parada desde Panel MS050
      ParadaPanelMS051 : Bool;   // Parada desde Panel MS051
      ParadaPanelMS052 : Bool;   // Parada desde Panel MS052
      ParadaPanelMS053 : Bool;   // Parada desde Panel MS053
      HabMS050 : Bool;   // Habilitado MS050
      HabMS051 : Bool;   // Habilitado MS051
      HabMS052 : Bool;   // Habilitado MS052
      HabMS053 : Bool;   // Habilitado MS053
      DeshabMS050 : Bool;   // Deshabilitado MS050
      DeshabMS051 : Bool;   // Deshabilitado MS051
      DeshabMS052 : Bool;   // Deshabilitado MS052
      DeshabMS053 : Bool;   // Deshabilitado MS053
      MarchaMS050 : Bool;   // Marchando MS050
      MarchaMS051 : Bool;   // Marchando MS051
      MarchaMS052 : Bool;   // Marchando MS052
      MarchaMS053 : Bool;   // Marchando MS053
      ParadaMS050 : Bool;   // Parando MS050
      ParadaMS051 : Bool;   // Parando MS051
      ParadaMS052 : Bool;   // Parando MS052
      ParadaMS053 : Bool;   // Parando MS053
      AnimMS050 : Byte;   // Animación MS050
      AnimMS051 : Byte;   // Animación MS051
      AnimMS052 : Byte;   // Animación MS052
      AnimMS053 : Byte;   // Animación MS053
      FallaGMTMS050 : Bool;   // Falla Térmica MS050
      FallaGMTMS051 : Bool;   // Falla Térmica MS051
      FallaGMTMS052 : Bool;   // Falla Térmica MS052
      FallaGMTMS053 : Bool;   // Falla Térmica MS053
      FallaCTCMS050 : Bool;   // Falla Contactor MS050
      FallaCTCMS051 : Bool;   // Falla Contactor MS051
      FallaCTCMS052 : Bool;   // Falla Contactor MS052
      FallaCTCMS053 : Bool;   // Falla Contactor MS053
      MantMS050 : Bool;   // Mantenimiento MS050
      MantMS051 : Bool;   // Mantenimiento MS051
      MantMS052 : Bool;   // Mantenimiento MS052
      MantMS053 : Bool;   // Mantenimiento MS053
      Enc1MS050 : Int;   // Enclavamiento1 para Ms050
      Enc2MS050 : Int;   // Enclavamiento2 para Ms050
      Enc1MS051 : Int;   // Enclavamiento1 para Ms051
      Enc2MS051 : Int;   // Enclavamiento2 para Ms051
      Enc1MS052 : Int;   // Enclavamiento1 para Ms052
      Enc2MS052 : Int;   // Enclavamiento2 para Ms052
      Enc1MS053 : Int;   // Enclavamiento1 para Ms053
      Enc2MS053 : Int;   // Enclavamiento2 para Ms053
      AutoMS050 : Bool;   // Modo automático para MS050
      AutoMS051 : Bool;   // Modo automático para MS051
      AutoMS052 : Bool;   // Modo automático para MS052
      AutoMS053 : Bool;   // Modo automático para MS054
      AutoArrMS050 : Bool;   // Arranque automático MS050
      AutoArrMS051 : Bool;   // Arranque automático MS051
      AutoArrMS052 : Bool;   // Arranque automático MS052
      AutoArrMS053 : Bool;   // Arranque automático MS053
      Reserva2 : Bool;
      Reserva3 : Bool;
      Reserva4 : Bool;
      Reserva_15 : Bool;
      Reserva_16 : Bool;
      Reserva_17 : Bool;
      Reserva_18 : Bool;
      Reserva_19 : Bool;
      Reserva_110 : Bool;
      Reserva_111 : Bool;
      Reserva_112 : Bool;
      Reserva_113 : Bool;
      Reserva_114 : Bool;
      Reserva_115 : Bool;
      Reserva_116 : Bool;
      Reserva_117 : Bool;
      Reserva_118 : Bool;
      Reserva_119 : Bool;
      Reserva_120 : Bool;
      Reserva_121 : Bool;
      Reserva_122 : Bool;
      Reserva_123 : Bool;
      Reserva_124 : Bool;
      Reserva_125 : Bool;
      Reserva_126 : Bool;
      Reserva_127 : Bool;
      Reserva_128 : Bool;
      Reserva_129 : Bool;
      Reserva_130 : Bool;
      Reserva_131 : Bool;
      Reserva_132 : Bool;
      Reserva_133 : Bool;
      Reserva_134 : Bool;
      Reserva_135 : Bool;
      Reserva_136 : Bool;
      Reserva_137 : Bool;
      Reserva_138 : Bool;
      Reserva_139 : Bool;
      Reserva_140 : Bool;
      Reserva_141 : Bool;
      Reserva_142 : Bool;
      Reserva_143 : Bool;
   END_VAR
BEGIN
END_DATA_BLOCK

// folder: Secadores/Baja

DATA_BLOCK "PanelSecBaja"   // DB49
{ S7_Optimized_Access := 'FALSE' }
VERSION : 0.1
   VAR
      InhMS054 : Bool;   // Inhibición MS054
      InhMS055 : Bool;   // Inhibición MS055
      Flanco1MS054 : Bool;   // Flanco 1 MS054
      Flanco1MS055 : Bool;   // Flanco 1 MS055
      Flanco2MS054 : Bool;   // Flanco 2 MS054
      Flanco2MS055 : Bool;   // Flanco 2 MS055
      Flanco3MS054 : Bool;   // Flanco 3 MS054
      Flanco3MS055 : Bool;   // Flanco 3 MS055
      HabPanelMS054 : Bool;   // Habilitación desde Panel MS054
      HabPanelMS055 : Bool;   // Habilitación desde Panel MS055
      DeshabPanelMS054 : Bool;   // Deshabilitación desde Panel MS054
      DeshabPanelMS055 : Bool;   // Deshabilitación desde Panel MS055
      MarchaPanelMS054 : Bool;   // Marcha desde Panel MS054
      MarchaPanelMS055 : Bool;   // Marcha desde Panel MS055
      ParadaPanelMS054 : Bool;   // Parada desde Panel MS054
      ParadaPanelMS055 : Bool;   // Parada desde Panel MS055
      HabMS054 : Bool;   // Habilitado MS054
      HabMS055 : Bool;   // Habilitado MS055
      DeshabMS054 : Bool;   // Deshabilitado MS054
      DeshabMS055 : Bool;   // Deshabilitado MS055
      MarchaMS054 : Bool;   // Marchando MS054
      MarchaMS055 : Bool;   // Marchando MS055
      ParadaMS054 : Bool;   // Parando MS054
      ParadaMS055 : Bool;   // Parando MS055
      AnimMS054 : Byte;   // Animación MS054
      AnimMS055 : Byte;   // Animación MS055
      FallaGMTMS054 : Bool;   // Falla Térmica MS054
      FallaGMTMS055 : Bool;   // Falla Térmica MS055
      FallaCTCMS054 : Bool;   // Falla Contactor MS054
      FallaCTCMS055 : Bool;   // Falla Contactor MS055
      MantMS054 : Bool;   // Mantenimiento MS054
      MantMS055 : Bool;   // Mantenimiento MS055
      Reserva2 : Bool;
      Reserva3 : Bool;
      Reserva4 : Bool;
      Reserva_15 : Bool;
      Reserva_16 : Bool;
      Reserva_17 : Bool;
      Reserva_18 : Bool;
      Reserva_19 : Bool;
      Reserva_110 : Bool;
      Reserva_111 : Bool;
      Reserva_112 : Bool;
      Reserva_113 : Bool;
      Reserva_114 : Bool;
      Reserva_115 : Bool;
      Reserva_116 : Bool;
      Reserva_117 : Bool;
      Reserva_118 : Bool;
      Reserva_119 : Bool;
      Reserva_120 : Bool;
      Reserva_121 : Bool;
      Reserva_122 : Bool;
      Reserva_123 : Bool;
      Reserva_124 : Bool;
      Reserva_125 : Bool;
      Reserva_126 : Bool;
      Reserva_127 : Bool;
      Reserva_128 : Bool;
      Reserva_129 : Bool;
      Reserva_130 : Bool;
      Reserva_131 : Bool;
      Reserva_132 : Bool;
      Reserva_133 : Bool;
      Reserva_134 : Bool;
      Reserva_135 : Bool;
      Reserva_136 : Bool;
      Reserva_137 : Bool;
      Reserva_138 : Bool;
      Reserva_139 : Bool;
      Reserva_140 : Bool;
      Reserva_141 : Bool;
      Reserva_142 : Bool;
      Reserva_143 : Bool;
   END_VAR
BEGIN
END_DATA_BLOCK

// folder: Torres de Agua/Torres Cavaleto

